         END_STRUCT;
         Reserve_5 : Struct
            ER_465 : Bool;   // Reserve
            ER_466 : Bool;   // Reserve
            ER_467 : Bool;   // Reserve
            ER_468 : Bool;   // Reserve
            ER_469 : Bool;   // Reserve
            ER_470 : Bool;   // Reserve
            ER_471 : Bool;   // Reserve
            ER_472 : Bool;   // Reserve
            ER_473 : Bool;   // Reserve
            ER_474 : Bool;   // Reserve
            ER_475 : Bool;   // Reserve
            ER_476 : Bool;   // Reserve
            ER_477 : Bool;   // Reserve
            ER_478 : Bool;   // Reserve
            ER_479 : Bool;   // Reserve
            ER_480 : Bool;   // Reserve
         END_STRUCT;
         Reserve_6 : Struct   // Meldungen Reserve
            ER_301 : Bool;   // Reserve
            ER_302 : Bool;   // Reserve
            ER_303 : Bool;   // Reserve
            ER_304 : Bool;   // Reserve
            ER_305 : Bool;   // Reserve
            ER_306 : Bool;   // Reserve
            ER_307 : Bool;   // Reserve
            ER_308 : Bool;   // Reserve
            ER_309 : Bool;   // Reserve
            ER_310 : Bool;   // Reserve
            ER_311 : Bool;   // Reserve
            ER_312 : Bool;   // Reserve
            ER_313 : Bool;   // Reserve
            ER_314 : Bool;   // Reserve
            ER_315 : Bool;   // Reserve
            ER_316 : Bool;   // Reserve
         END_STRUCT;
         Reserve_7 : Struct   // Meldungen Reserve
            ER_317 : Bool;   // Reserve
            ER_318 : Bool;   // Reserve
            ER_319 : Bool;   // Reserve
            ER_320 : Bool;   // Reserve
            ER_321 : Bool;   // Reserve
            ER_322 : Bool;   // Reserve
            ER_323 : Bool;   // Reserve
            ER_324 : Bool;   // Reserve
            ER_325 : Bool;   // Reserve
            ER_326 : Bool;   // Reserve
            ER_327 : Bool;   // Reserve
            ER_328 : Bool;   // Reserve
            ER_329 : Bool;   // Reserve
            ER_330 : Bool;   // Reserve
            ER_331 : Bool;   // Reserve
            ER_332 : Bool;   // Reserve
         END_STRUCT;
         Reserve_8 : Struct   // FU Reserve
            ER_333 : Bool;   // Störung Reserve FU 1: Überstrom
            ER_334 : Bool;   // Störung Reserve FU 1: Zwischenkreisspannung Überspannung
            ER_335 : Bool;   // Störung Reserve FU 1: Zwischenkreisspannung Unterspannung
            ER_336 : Bool;   // Störung Reserve FU 1: Übertemperatur Kühlkörper Wechselrichter
            ER_337 : Bool;   // Störung Reserve FU 1: Motordatenidentifikation fehlerhaft
            ER_338 : Bool;   // Störung Reserve FU 1: Erdschluss
            ER_339 : Bool;   // Störung Reserve FU 1: Reserve
            ER_340 : Bool;   // Störung Reserve FU 1: Führung durch PLC fehlt
            ER_341 : Bool;   // Störung Reserve FU 1: Reserve
            ER_342 : Bool;   // Störung Reserve FU 1: Reserve
            ER_343 : Bool;   // Störung Reserve FU 1: Reserve
            ER_344_ : Bool;   // Störung Reserve FU 1: Reserve
            ER_345 : Bool;   // Störung Reserve FU 1: Reserve
            ER_346 : Bool;   // Störung Reserve FU 1: Reserve
            ER_347 : Bool;   // Störung Reserve FU 1: Reserve
            ER_348 : Bool;   // Störung Reserve FU 1: Reserve
         END_STRUCT;
         Reserve_9 : Struct
            ER_349 : Bool;   // Reserve
            ER_350 : Bool;   // Reserve
            ER_351 : Bool;   // Reserve
            ER_352 : Bool;   // Reserve
            ER_353 : Bool;   // Reserve
            ER_354 : Bool;   // Reserve
            ER_355 : Bool;   // Reserve
            ER_356 : Bool;   // Reserve
            ER_357 : Bool;   // Reserve
            ER_358 : Bool;   // Reserve
            ER_359 : Bool;   // Reserve
            ER_360 : Bool;   // Reserve
            ER_361 : Bool;   // Reserve
            ER_362 : Bool;   // Reserve
            ER_363 : Bool;   // Reserve
            ER_364 : Bool;   // Reserve
         END_STRUCT;
         Reserve_10 : Struct   // FU Reserve
            ER_365 : Bool;   // Störung Reserve FU 2: Überstrom
            ER_366 : Bool;   // Störung Reserve FU 2: Zwischenkreisspannung Überspannung
            ER_367 : Bool;   // Störung Reserve FU 2: Zwischenkreisspannung Unterspannung
            ER_368 : Bool;   // Störung Reserve FU 2: Übertemperatur Kühlkörper Wechselrichter
            ER_369 : Bool;   // Störung Reserve FU 2: Motordatenidentifikation fehlerhaft
            ER_370 : Bool;   // Störung Reserve FU 2: Erdschluss
            ER_371 : Bool;   // Störung Reserve FU 2: Reserve
            ER_372 : Bool;   // Störung Reserve FU 2: Führung durch PLC fehlt
            ER_373 : Bool;   // Störung Reserve FU 2: Reserve
            ER_374 : Bool;   // Störung Reserve FU 2: Reserve
            ER_375 : Bool;   // Störung Reserve FU 2: Reserve
            ER_376 : Bool;   // Störung Reserve FU 2: Reserve
            ER_377 : Bool;   // Störung Reserve FU 2: Reserve
            ER_378 : Bool;   // Störung Reserve FU 2: Reserve
            ER_379 : Bool;   // Störung Reserve FU 2: Reserve
            ER_380 : Bool;   // Störung Reserve FU 2: Reserve
         END_STRUCT;
         SDC : Struct   // SDC Störungs
            ER_901 : Bool;   // Reserve
            ER_902 : Bool;   // Reserve
            ER_903 : Bool;   // Störung SDC Positionssprung
            ER_904 : Bool;   // Störung SDC keine Sektion gefunden
            ER_905 : Bool;   // Störung SDC Kommandos nicht plausibel
            ER_906 : Bool;   // Störung SDC Positionsgrenzen
            ER_907 : Bool;   // Störung SDC falsche EMS Nummer
            ER_908 : Bool;   // Störung SDC falsche Sektion Nummer
            ER_909 : Bool;   // Reserve
            ER_910 : Bool;   // Reserve
            ER_911 : Bool;   // Reserve
            ER_912 : Bool;   // Reserve
            ER_913 : Bool;   // Reserve
            ER_914 : Bool;   // Reserve
            ER_915 : Bool;   // Reserve
            ER_916 : Bool;   // Reserve
         END_STRUCT;
      END_STRUCT;
      EMS_ER_WORDs : Array[1..200] of Struct   // EMS Störung WORDs
         ER_WORD : Array[0..24] of Word;   // Störworte
      END_STRUCT;
      SDC : Struct
         ER_917 : Bool;   // Störung SDC Kommunikation mit Anlagensteuerung
         ER_918 : Bool;   // Störung SDC Safety Kommunikation mit Anlagensteuerung
         ER_919 : Bool;   // Störung SDC Reserve
         ER_920 : Bool;   // Störung SDC Reserve
         ER_921 : Bool;   // Störung SDC Reserve
         ER_922 : Bool;   // Störung SDC Reserve
         ER_923 : Bool;   // Störung SDC Reserve
         ER_924 : Bool;   // Störung SDC Reserve
         ER_925 : Bool;   // Störung SDC OB80 Zykluszeit
         ER_926 : Bool;   // Störung SDC OB82 Diagnosealarm
         ER_927 : Bool;   // Störung SDC OB83 Baugruppenwechsel
         ER_928 : Bool;   // Störung SDC OB86 Baugruppenträger ausgefallen
         ER_929 : Bool;   // Störung SDC OB121 Programmierfehler
         ER_930 : Bool;   // Störung SDC OB122 Peripherie-Zugriff
         ER_931 : Bool;   // Störung SDC Reserve
         ER_932 : Bool;   // Störung SDC Reserve
      END_STRUCT;
   END_VAR
BEGIN
END_DATA_BLOCK

DATA_BLOCK "DB_SDC_ERRORS_STAT"   // DB3724
{ S7_Optimized_Access := 'FALSE' }
VERSION : 0.1
   VAR
      HEADER : Struct   // Struktur für Datenheader // nicht verschieben
         DB_NR : Int := 3724;   // DB Nummer
         MIN_NR_FAULT_STAT : Int := 1;   // Niedrigste Fehler Nummer im Daten DB
         MAX_NR_FAULT_STAT : Int := 200;   // Höchste Fehler Nummer im Daten DB
         START_FAULT_STAT : Int := 20;   // Startadresse der Fehler Daten im Daten DB
         LAENGE_FAULT_STAT : Int := 28;   // Länge Fehler Daten
         FAULT_PRO_SEITE_HMI : Int := 10;   // Reserve
         RES12 : Int := 0;   // Reserve
         RES14 : Int := 0;   // Reserve
         RES16 : Int := 0;   // Reserve
         LOAD : Bool := FALSE;   // "0" zum laden des DB auf CPU
         RESET_ARCH : Bool := FALSE;   // Archiv löschen
      END_STRUCT;
      ER_ARCHIV : Array[1..1000] of "UDT_SDC_ERROR_STAT";   // Error Archiv
      ER_AKT : Array[1..200] of Struct   // Error aktiv EMS
         ER_TRIGER : Word;   // Error auslösen Aktiv von EMS
         ER_STAT : Array[1..4] of "UDT_SDC_TS_IF_STATUS_VAL";   // Error Status Aktiv EMS
      END_STRUCT;
   END_VAR
BEGIN
   ER_ARCHIV[1].EMS_TS_STAT_VAL.EMS_ID := 0;
   ER_ARCHIV[1].EMS_TS_STAT_VAL.PROFIL := 0;
   ER_ARCHIV[1].EMS_TS_STAT_VAL.DRIVE_POS := 0;
   ER_ARCHIV[1].EMS_TS_STAT_VAL.HOIST_POS := 0;
   ER_ARCHIV[1].EMS_TS_STAT_VAL.ERROR := 0;
   ER_ARCHIV[1].EMS_TS_STAT_VAL.DRIVE_POS_PERC := 0;
   ER_ARCHIV[1].EMS_TS_STAT_VAL.SEK := 0;
   ER_ARCHIV[1].ER._901_ER_SUM := FALSE;
   ER_ARCHIV[1].ER._902_ER_SUM_SDC := FALSE;
   ER_ARCHIV[1].ER._903_ER_BC_JUMP := FALSE;
   ER_ARCHIV[1].ER._904_ER_NO_SEK := FALSE;
   ER_ARCHIV[1].ER._905_ER_COMMAND := FALSE;
   ER_ARCHIV[1].ER._906_ER_BC_LIM := FALSE;
   ER_ARCHIV[1].ER._907_ER_EMS_ID := FALSE;
   ER_ARCHIV[1].ER._908_ER_SEK_NR := FALSE;
   ER_ARCHIV[1].ER._909_ER_LIFE := FALSE;
   ER_ARCHIV[1].ER._910_ER_BUS := FALSE;
   ER_ARCHIV[1].ER._911 := FALSE;
   ER_ARCHIV[1].ER._912 := FALSE;
   ER_ARCHIV[1].ER._913 := FALSE;
   ER_ARCHIV[1].ER._914 := FALSE;
   ER_ARCHIV[1].ER._915 := FALSE;
   ER_ARCHIV[1].ER._916 := FALSE;
   ER_ARCHIV[1].Spare := 0;
   ER_ARCHIV[1].ER_DATE := DT#1990-01-01-00:00:00;
   ER_ARCHIV[2].EMS_TS_STAT_VAL.EMS_ID := 0;
   ER_ARCHIV[2].EMS_TS_STAT_VAL.PROFIL := 0;
   ER_ARCHIV[2].EMS_TS_STAT_VAL.DRIVE_POS := 0;
   ER_ARCHIV[2].EMS_TS_STAT_VAL.HOIST_POS := 0;
   ER_ARCHIV[2].EMS_TS_STAT_VAL.ERROR := 0;
   ER_ARCHIV[2].EMS_TS_STAT_VAL.DRIVE_POS_PERC := 0;
   ER_ARCHIV[2].EMS_TS_STAT_VAL.SEK := 0;
   ER_ARCHIV[2].ER._901_ER_SUM := FALSE;
   ER_ARCHIV[2].ER._902_ER_SUM_SDC := FALSE;
   ER_ARCHIV[2].ER._903_ER_BC_JUMP := FALSE;
   ER_ARCHIV[2].ER._904_ER_NO_SEK := FALSE;
   ER_ARCHIV[2].ER._905_ER_COMMAND := FALSE;
   ER_ARCHIV[2].ER._906_ER_BC_LIM := FALSE;
   ER_ARCHIV[2].ER._907_ER_EMS_ID := FALSE;
   ER_ARCHIV[2].ER._908_ER_SEK_NR := FALSE;
   ER_ARCHIV[2].ER._909_ER_LIFE := FALSE;
   ER_ARCHIV[2].ER._910_ER_BUS := FALSE;
   ER_ARCHIV[2].ER._911 := FALSE;
   ER_ARCHIV[2].ER._912 := FALSE;
   ER_ARCHIV[2].ER._913 := FALSE;
   ER_ARCHIV[2].ER._914 := FALSE;
   ER_ARCHIV[2].ER._915 := FALSE;
   ER_ARCHIV[2].ER._916 := FALSE;
   ER_ARCHIV[2].Spare := 0;
   ER_ARCHIV[2].ER_DATE := DT#1990-01-01-00:00:00;
   ER_ARCHIV[3].EMS_TS_STAT_VAL.EMS_ID := 0;
   ER_ARCHIV[3].EMS_TS_STAT_VAL.PROFIL := 0;
   ER_ARCHIV[3].EMS_TS_STAT_VAL.DRIVE_POS := 0;
   ER_ARCHIV[3].EMS_TS_STAT_VAL.HOIST_POS := 0;
   ER_ARCHIV[3].EMS_TS_STAT_VAL.ERROR := 0;
   ER_ARCHIV[3].EMS_TS_STAT_VAL.DRIVE_POS_PERC := 0;
   ER_ARCHIV[3].EMS_TS_STAT_VAL.SEK := 0;
   ER_ARCHIV[3].ER._901_ER_SUM := FALSE;
   ER_ARCHIV[3].ER._902_ER_SUM_SDC := FALSE;
   ER_ARCHIV[3].ER._903_ER_BC_JUMP := FALSE;
   ER_ARCHIV[3].ER._904_ER_NO_SEK := FALSE;
   ER_ARCHIV[3].ER._905_ER_COMMAND := FALSE;
   ER_ARCHIV[3].ER._906_ER_BC_LIM := FALSE;
   ER_ARCHIV[3].ER._907_ER_EMS_ID := FALSE;
   ER_ARCHIV[3].ER._908_ER_SEK_NR := FALSE;
   ER_ARCHIV[3].ER._909_ER_LIFE := FALSE;
   ER_ARCHIV[3].ER._910_ER_BUS := FALSE;
   ER_ARCHIV[3].ER._911 := FALSE;
   ER_ARCHIV[3].ER._912 := FALSE;
   ER_ARCHIV[3].ER._913 := FALSE;
   ER_ARCHIV[3].ER._914 := FALSE;
   ER_ARCHIV[3].ER._915 := FALSE;
   ER_ARCHIV[3].ER._916 := FALSE;
   ER_ARCHIV[3].Spare := 0;
   ER_ARCHIV[3].ER_DATE := DT#1990-01-01-00:00:00;
   ER_ARCHIV[4].EMS_TS_STAT_VAL.EMS_ID := 0;
   ER_ARCHIV[4].EMS_TS_STAT_VAL.PROFIL := 0;
   ER_ARCHIV[4].EMS_TS_STAT_VAL.DRIVE_POS := 0;
   ER_ARCHIV[4].EMS_TS_STAT_VAL.HOIST_POS := 0;
   ER_ARCHIV[4].EMS_TS_STAT_VAL.ERROR := 0;
   ER_ARCHIV[4].EMS_TS_STAT_VAL.DRIVE_POS_PERC := 0;
   ER_ARCHIV[4].EMS_TS_STAT_VAL.SEK := 0;
   ER_ARCHIV[4].ER._901_ER_SUM := FALSE;
   ER_ARCHIV[4].ER._902_ER_SUM_SDC := FALSE;
   ER_ARCHIV[4].ER._903_ER_BC_JUMP := FALSE;
   ER_ARCHIV[4].ER._904_ER_NO_SEK := FALSE;
   ER_ARCHIV[4].ER._905_ER_COMMAND := FALSE;
   ER_ARCHIV[4].ER._906_ER_BC_LIM := FALSE;
   ER_ARCHIV[4].ER._907_ER_EMS_ID := FALSE;
   ER_ARCHIV[4].ER._908_ER_SEK_NR := FALSE;
   ER_ARCHIV[4].ER._909_ER_LIFE := FALSE;
   ER_ARCHIV[4].ER._910_ER_BUS := FALSE;
   ER_ARCHIV[4].ER._911 := FALSE;
   ER_ARCHIV[4].ER._912 := FALSE;
   ER_ARCHIV[4].ER._913 := FALSE;
   ER_ARCHIV[4].ER._914 := FALSE;
   ER_ARCHIV[4].ER._915 := FALSE;
   ER_ARCHIV[4].ER._916 := FALSE;
   ER_ARCHIV[4].Spare := 0;
   ER_ARCHIV[4].ER_DATE := DT#1990-01-01-00:00:00;
   ER_ARCHIV[5].EMS_TS_STAT_VAL.EMS_ID := 0;
   ER_ARCHIV[5].EMS_TS_STAT_VAL.PROFIL := 0;
   ER_ARCHIV[5].EMS_TS_STAT_VAL.DRIVE_POS := 0;
   ER_ARCHIV[5].EMS_TS_STAT_VAL.HOIST_POS := 0;
   ER_ARCHIV[5].EMS_TS_STAT_VAL.ERROR := 0;
   ER_ARCHIV[5].EMS_TS_STAT_VAL.DRIVE_POS_PERC := 0;
   ER_ARCHIV[5].EMS_TS_STAT_VAL.SEK := 0;
   ER_ARCHIV[5].ER._901_ER_SUM := FALSE;
   ER_ARCHIV[5].ER._902_ER_SUM_SDC := FALSE;
   ER_ARCHIV[5].ER._903_ER_BC_JUMP := FALSE;
   ER_ARCHIV[5].ER._904_ER_NO_SEK := FALSE;
   ER_ARCHIV[5].ER._905_ER_COMMAND := FALSE;
   ER_ARCHIV[5].ER._906_ER_BC_LIM := FALSE;
   ER_ARCHIV[5].ER._907_ER_EMS_ID := FALSE;
   ER_ARCHIV[5].ER._908_ER_SEK_NR := FALSE;
   ER_ARCHIV[5].ER._909_ER_LIFE := FALSE;
   ER_ARCHIV[5].ER._910_ER_BUS := FALSE;
   ER_ARCHIV[5].ER._911 := FALSE;
   ER_ARCHIV[5].ER._912 := FALSE;
   ER_ARCHIV[5].ER._913 := FALSE;
   ER_ARCHIV[5].ER._914 := FALSE;
   ER_ARCHIV[5].ER._915 := FALSE;
   ER_ARCHIV[5].ER._916 := FALSE;
   ER_ARCHIV[5].Spare := 0;
   ER_ARCHIV[5].ER_DATE := DT#1990-01-01-00:00:00;
   ER_ARCHIV[6].EMS_TS_STAT_VAL.EMS_ID := 0;
   ER_ARCHIV[6].EMS_TS_STAT_VAL.PROFIL := 0;
   ER_ARCHIV[6].EMS_TS_STAT_VAL.DRIVE_POS := 0;
   ER_ARCHIV[6].EMS_TS_STAT_VAL.HOIST_POS := 0;
   ER_ARCHIV[6].EMS_TS_STAT_VAL.ERROR := 0;
   ER_ARCHIV[6].EMS_TS_STAT_VAL.DRIVE_POS_PERC := 0;
   ER_ARCHIV[6].EMS_TS_STAT_VAL.SEK := 0;
   ER_ARCHIV[6].ER._901_ER_SUM := FALSE;
   ER_ARCHIV[6].ER._902_ER_SUM_SDC := FALSE;
   ER_ARCHIV[6].ER._903_ER_BC_JUMP := FALSE;
   ER_ARCHIV[6].ER._904_ER_NO_SEK := FALSE;
   ER_ARCHIV[6].ER._905_ER_COMMAND := FALSE;
   ER_ARCHIV[6].ER._906_ER_BC_LIM := FALSE;
   ER_ARCHIV[6].ER._907_ER_EMS_ID := FALSE;
   ER_ARCHIV[6].ER._908_ER_SEK_NR := FALSE;
   ER_ARCHIV[6].ER._909_ER_LIFE := FALSE;
   ER_ARCHIV[6].ER._910_ER_BUS := FALSE;
   ER_ARCHIV[6].ER._911 := FALSE;
   ER_ARCHIV[6].ER._912 := FALSE;
   ER_ARCHIV[6].ER._913 := FALSE;
   ER_ARCHIV[6].ER._914 := FALSE;
   ER_ARCHIV[6].ER._915 := FALSE;
   ER_ARCHIV[6].ER._916 := FALSE;
   ER_ARCHIV[6].Spare := 0;
   ER_ARCHIV[6].ER_DATE := DT#1990-01-01-00:00:00;
   ER_ARCHIV[7].EMS_TS_STAT_VAL.EMS_ID := 0;
   ER_ARCHIV[7].EMS_TS_STAT_VAL.PROFIL := 0;
   ER_ARCHIV[7].EMS_TS_STAT_VAL.DRIVE_POS := 0;
   ER_ARCHIV[7].EMS_TS_STAT_VAL.HOIST_POS := 0;
   ER_ARCHIV[7].EMS_TS_STAT_VAL.ERROR := 0;
   ER_ARCHIV[7].EMS_TS_STAT_VAL.DRIVE_POS_PERC := 0;
   ER_ARCHIV[7].EMS_TS_STAT_VAL.SEK := 0;
   ER_ARCHIV[7].ER._901_ER_SUM := FALSE;
   ER_ARCHIV[7].ER._902_ER_SUM_SDC := FALSE;
   ER_ARCHIV[7].ER._903_ER_BC_JUMP := FALSE;
   ER_ARCHIV[7].ER._904_ER_NO_SEK := FALSE;
   ER_ARCHIV[7].ER._905_ER_COMMAND := FALSE;
   ER_ARCHIV[7].ER._906_ER_BC_LIM := FALSE;
   ER_ARCHIV[7].ER._907_ER_EMS_ID := FALSE;
   ER_ARCHIV[7].ER._908_ER_SEK_NR := FALSE;
   ER_ARCHIV[7].ER._909_ER_LIFE := FALSE;
   ER_ARCHIV[7].ER._910_ER_BUS := FALSE;
   ER_ARCHIV[7].ER._911 := FALSE;
   ER_ARCHIV[7].ER._912 := FALSE;
   ER_ARCHIV[7].ER._913 := FALSE;
   ER_ARCHIV[7].ER._914 := FALSE;
   ER_ARCHIV[7].ER._915 := FALSE;
   ER_ARCHIV[7].ER._916 := FALSE;
   ER_ARCHIV[7].Spare := 0;
   ER_ARCHIV[7].ER_DATE := DT#1990-01-01-00:00:00;
   ER_ARCHIV[8].EMS_TS_STAT_VAL.EMS_ID := 0;
   ER_ARCHIV[8].EMS_TS_STAT_VAL.PROFIL := 0;
   ER_ARCHIV[8].EMS_TS_STAT_VAL.DRIVE_POS := 0;
   ER_ARCHIV[8].EMS_TS_STAT_VAL.HOIST_POS := 0;
   ER_ARCHIV[8].EMS_TS_STAT_VAL.ERROR := 0;
   ER_ARCHIV[8].EMS_TS_STAT_VAL.DRIVE_POS_PERC := 0;
   ER_ARCHIV[8].EMS_TS_STAT_VAL.SEK := 0;
   ER_ARCHIV[8].ER._901_ER_SUM := FALSE;
   ER_ARCHIV[8].ER._902_ER_SUM_SDC := FALSE;
   ER_ARCHIV[8].ER._903_ER_BC_JUMP := FALSE;
   ER_ARCHIV[8].ER._904_ER_NO_SEK := FALSE;
   ER_ARCHIV[8].ER._905_ER_COMMAND := FALSE;
   ER_ARCHIV[8].ER._906_ER_BC_LIM := FALSE;
   ER_ARCHIV[8].ER._907_ER_EMS_ID := FALSE;
   ER_ARCHIV[8].ER._908_ER_SEK_NR := FALSE;
   ER_ARCHIV[8].ER._909_ER_LIFE := FALSE;
   ER_ARCHIV[8].ER._910_ER_BUS := FALSE;
   ER_ARCHIV[8].ER._911 := FALSE;
   ER_ARCHIV[8].ER._912 := FALSE;
   ER_ARCHIV[8].ER._913 := FALSE;
   ER_ARCHIV[8].ER._914 := FALSE;
   ER_ARCHIV[8].ER._915 := FALSE;
   ER_ARCHIV[8].ER._916 := FALSE;
   ER_ARCHIV[8].Spare := 0;
   ER_ARCHIV[8].ER_DATE := DT#1990-01-01-00:00:00;
   // 30600 more start values not shown
END_DATA_BLOCK

DATA_BLOCK "DB_SDC_EMS_SIM"   // DB3726
{ S7_Optimized_Access := 'FALSE' }
VERSION : 0.1
   VAR
      HEADER : Struct   // Struktur für Datenheader // nicht verschieben
         DB_NR : Int := 3726;   // DB Nummer
         MIN_NR_EMS : Int := 1;   // Niedrigste EMS Nummer im Daten DB
         MAX_NR_EMS : Int := 200;   // Höchste EMS Nummer im Daten DB
         START_DAT : Int := 40;   // Startadresse der EMS Daten im Daten DB
         LAENGE_EMS : Int := 40;   // Länge Eingänge pro EMS
         RES10 : Int := 0;   // Reserve
         RES12 : Int := 0;   // Reserve
         RES14 : Int := 0;   // Reserve
         RES16 : Int := 0;   // Reserve
         RES18 : Int := 0;   // Reserve
      END_STRUCT;
      PAR : Struct   // Parameter Simulation
         BARCODE_START : DInt := 1;   // min Barcodevalue
         BARCODE_ENDE : DInt := 500000;   // max Barcodevalue
         HUB_START : Int := 0;   // min Hoistvalue
         HUB_ENDE : Int := 4010;   // max Hoistvalue
         LEAP_AKT : Array[1..20] of Bool;   // Leap Aktiv
         LEAP_HIGH_LOW : Array[1..20] of Bool;   // Leap Aktiv
         ON : Bool := TRUE;   // Simulation ON "1"
         RES18 : Int := 0;   // Reserve
      END_STRUCT;
      EMS : Array[1..200] of "UDT_EMS_IF_Q";   // EMS Simulation Eingänge
      EMS_TEMP : "UDT_EMS_IF_Q";
   END_VAR
BEGIN
   PAR.LEAP_AKT[1] := TRUE;
   PAR.LEAP_AKT[2] := TRUE;
   PAR.LEAP_AKT[3] := TRUE;
   PAR.LEAP_HIGH_LOW[1] := TRUE;
   PAR.LEAP_HIGH_LOW[2] := FALSE;
   PAR.LEAP_HIGH_LOW[3] := TRUE;
   PAR.LEAP_AKT[4] := FALSE;
   PAR.LEAP_AKT[5] := FALSE;
   PAR.LEAP_AKT[6] := FALSE;
   PAR.LEAP_AKT[7] := FALSE;
   PAR.LEAP_AKT[8] := FALSE;
   PAR.LEAP_AKT[9] := FALSE;
   PAR.LEAP_AKT[10] := FALSE;
   PAR.LEAP_AKT[11] := FALSE;
   PAR.LEAP_AKT[12] := FALSE;
   PAR.LEAP_AKT[13] := FALSE;
   PAR.LEAP_AKT[14] := FALSE;
   PAR.LEAP_AKT[15] := FALSE;
   PAR.LEAP_AKT[16] := FALSE;
   PAR.LEAP_AKT[17] := FALSE;
   PAR.LEAP_AKT[18] := FALSE;
   PAR.LEAP_AKT[19] := FALSE;
   PAR.LEAP_AKT[20] := FALSE;
   PAR.LEAP_HIGH_LOW[4] := FALSE;
   PAR.LEAP_HIGH_LOW[5] := FALSE;
   PAR.LEAP_HIGH_LOW[6] := FALSE;
   PAR.LEAP_HIGH_LOW[7] := FALSE;
   PAR.LEAP_HIGH_LOW[8] := FALSE;
   PAR.LEAP_HIGH_LOW[9] := FALSE;
   PAR.LEAP_HIGH_LOW[10] := FALSE;
   PAR.LEAP_HIGH_LOW[11] := FALSE;
   PAR.LEAP_HIGH_LOW[12] := FALSE;
   PAR.LEAP_HIGH_LOW[13] := FALSE;
   PAR.LEAP_HIGH_LOW[14] := FALSE;
   PAR.LEAP_HIGH_LOW[15] := FALSE;
   PAR.LEAP_HIGH_LOW[16] := FALSE;
   PAR.LEAP_HIGH_LOW[17] := FALSE;
   PAR.LEAP_HIGH_LOW[18] := FALSE;
   PAR.LEAP_HIGH_LOW[19] := FALSE;
   PAR.LEAP_HIGH_LOW[20] := FALSE;
   EMS[1].STAT.LIFE_BIT := TRUE;
   EMS[1].STAT.ER_SUM := FALSE;
   EMS[1].STAT.IR_MAN := FALSE;
   EMS[1].STAT.ER_RESET := FALSE;
   EMS[1].STAT.HOIST_CLEAR := FALSE;
   EMS[1].STAT.POS_START_X := FALSE;
   EMS[1].STAT.ALWAYS_ONE := TRUE;
   EMS[1].STAT.H_DISABLED := FALSE;
   EMS[1].STAT.D_FWD := TRUE;
   EMS[1].STAT.D_RWD := FALSE;
   EMS[1].STAT.bit12 := FALSE;
   EMS[1].STAT.D_IN_POS := FALSE;
   EMS[1].STAT.H_UP := FALSE;
   EMS[1].STAT.H_DOWN := FALSE;
   EMS[1].STAT.H_IN_POS := TRUE;
   EMS[1].STAT.H_IN_TOPPOS := FALSE;
   EMS[1].STAT.bit2_0 := FALSE;
   EMS[1].STAT.bit2_1 := FALSE;
   EMS[1].STAT.bit2_2 := FALSE;
   EMS[1].STAT.bit2_3 := FALSE;
   EMS[1].STAT.IN_BOTPOS := FALSE;
   EMS[1].STAT.bit2_5 := FALSE;
   EMS[1].STAT.bit2_6 := FALSE;
   EMS[1].STAT.bit2_7 := FALSE;
   EMS[1].STAT.MESS_POS := FALSE;
   EMS[1].STAT.bit3_2 := FALSE;
   EMS[1].STAT.bit3_3 := FALSE;
   EMS[1].STAT.bit3_4 := FALSE;
   EMS[1].STAT.bit3_5 := FALSE;
   EMS[1].STAT.bit3_6 := FALSE;
   EMS[1].STAT.DATA_TRANS := FALSE;
   EMS[1].ERROR := 0;
   EMS[1].D_POS := 22899;
   EMS[1].H_POS := 603;
   EMS[1].ER_WORD_No := 1;
   EMS[1].ER_WORD := 16#0000;
   EMS[1].FB_DBNo := 0;
   EMS[1].FB_DBBNo := 0;
   EMS[2].STAT.LIFE_BIT := TRUE;
   EMS[2].STAT.ER_SUM := FALSE;
   EMS[2].STAT.IR_MAN := FALSE;
   EMS[2].STAT.ER_RESET := FALSE;
   EMS[2].STAT.HOIST_CLEAR := FALSE;
   EMS[2].STAT.POS_START_X := FALSE;
   EMS[2].STAT.ALWAYS_ONE := TRUE;
   EMS[2].STAT.H_DISABLED := FALSE;
   EMS[2].STAT.D_FWD := TRUE;
   EMS[2].STAT.D_RWD := FALSE;
   EMS[2].STAT.bit12 := FALSE;
   EMS[2].STAT.D_IN_POS := FALSE;
   EMS[2].STAT.H_UP := FALSE;
   EMS[2].STAT.H_DOWN := FALSE;
   EMS[2].STAT.H_IN_POS := FALSE;
   EMS[2].STAT.H_IN_TOPPOS := TRUE;
   EMS[2].STAT.bit2_0 := FALSE;
   EMS[2].STAT.bit2_1 := FALSE;
   EMS[2].STAT.bit2_2 := FALSE;
   EMS[2].STAT.bit2_3 := FALSE;
   EMS[2].STAT.IN_BOTPOS := FALSE;
   EMS[2].STAT.bit2_5 := FALSE;
   EMS[2].STAT.bit2_6 := FALSE;
   EMS[2].STAT.bit2_7 := FALSE;
   EMS[2].STAT.MESS_POS := FALSE;
   EMS[2].STAT.bit3_2 := FALSE;
   EMS[2].STAT.bit3_3 := FALSE;
   EMS[2].STAT.bit3_4 := FALSE;
   EMS[2].STAT.bit3_5 := FALSE;
   EMS[2].STAT.bit3_6 := FALSE;
   EMS[2].STAT.DATA_TRANS := FALSE;
   EMS[2].ERROR := 0;
   EMS[2].D_POS := 10522;
   EMS[2].H_POS := 4010;
   EMS[2].ER_WORD_No := 1;
   EMS[2].ER_WORD := 16#0000;
   EMS[2].FB_DBNo := 0;
   EMS[2].FB_DBBNo := 0;
   EMS[3].STAT.LIFE_BIT := TRUE;
   EMS[3].STAT.ER_SUM := FALSE;
   EMS[3].STAT.IR_MAN := FALSE;
   EMS[3].STAT.ER_RESET := FALSE;
   EMS[3].STAT.HOIST_CLEAR := FALSE;
   EMS[3].STAT.POS_START_X := FALSE;
   EMS[3].STAT.ALWAYS_ONE := TRUE;
   EMS[3].STAT.H_DISABLED := FALSE;
   EMS[3].STAT.D_FWD := TRUE;
   EMS[3].STAT.D_RWD := FALSE;
   EMS[3].STAT.bit12 := FALSE;
   EMS[3].STAT.D_IN_POS := FALSE;
   EMS[3].STAT.H_UP := FALSE;
   EMS[3].STAT.H_DOWN := FALSE;
   EMS[3].STAT.H_IN_POS := FALSE;
   EMS[3].STAT.H_IN_TOPPOS := TRUE;
   EMS[3].STAT.bit2_0 := FALSE;
   EMS[3].STAT.bit2_1 := FALSE;
   EMS[3].STAT.bit2_2 := FALSE;
   EMS[3].STAT.bit2_3 := FALSE;
   EMS[3].STAT.IN_BOTPOS := FALSE;
   EMS[3].STAT.bit2_5 := FALSE;
   EMS[3].STAT.bit2_6 := FALSE;
   EMS[3].STAT.bit2_7 := FALSE;
   EMS[3].STAT.MESS_POS := FALSE;
   EMS[3].STAT.bit3_2 := FALSE;
   EMS[3].STAT.bit3_3 := FALSE;
   EMS[3].STAT.bit3_4 := FALSE;
   EMS[3].STAT.bit3_5 := FALSE;
   EMS[3].STAT.bit3_6 := FALSE;
   EMS[3].STAT.DATA_TRANS := FALSE;
   EMS[3].ERROR := 0;
   EMS[3].D_POS := 96650;
   EMS[3].H_POS := 4010;
   EMS[3].ER_WORD_No := 1;
   EMS[3].ER_WORD := 16#0000;
   EMS[3].FB_DBNo := 0;
   EMS[3].FB_DBBNo := 0;
   EMS[4].STAT.LIFE_BIT := FALSE;
   EMS[4].STAT.ER_SUM := FALSE;
   EMS[4].STAT.IR_MAN := FALSE;
   EMS[4].STAT.ER_RESET := FALSE;
   EMS[4].STAT.HOIST_CLEAR := FALSE;
   EMS[4].STAT.POS_START_X := FALSE;
   EMS[4].STAT.ALWAYS_ONE := FALSE;
   EMS[4].STAT.H_DISABLED := FALSE;
   EMS[4].STAT.D_FWD := FALSE;
   EMS[4].STAT.D_RWD := FALSE;
   EMS[4].STAT.bit12 := FALSE;
   EMS[4].STAT.D_IN_POS := FALSE;
   EMS[4].STAT.H_UP := FALSE;
   EMS[4].STAT.H_DOWN := FALSE;
   EMS[4].STAT.H_IN_POS := FALSE;
   EMS[4].STAT.H_IN_TOPPOS := FALSE;
   EMS[4].STAT.bit2_0 := FALSE;
   EMS[4].STAT.bit2_1 := FALSE;
   EMS[4].STAT.bit2_2 := FALSE;
   EMS[4].STAT.bit2_3 := FALSE;
   EMS[4].STAT.IN_BOTPOS := FALSE;
   EMS[4].STAT.bit2_5 := FALSE;
   EMS[4].STAT.bit2_6 := FALSE;
   EMS[4].STAT.bit2_7 := FALSE;
   EMS[4].STAT.MESS_POS := FALSE;
   EMS[4].STAT.bit3_2 := FALSE;
   EMS[4].STAT.bit3_3 := FALSE;
   EMS[4].STAT.bit3_4 := FALSE;
   EMS[4].STAT.bit3_5 := FALSE;
   EMS[4].STAT.bit3_6 := FALSE;
   EMS[4].STAT.DATA_TRANS := FALSE;
   EMS[4].ERROR := 0;
   EMS[4].D_POS := 0;
   EMS[4].H_POS := 0;
   EMS[4].ER_WORD_No := 0;
   EMS[4].ER_WORD := 16#0000;
   EMS[4].FB_DBNo := 0;
   EMS[4].FB_DBBNo := 0;
   EMS[5].STAT.LIFE_BIT := FALSE;
   EMS[5].STAT.ER_SUM := FALSE;
   EMS[5].STAT.IR_MAN := FALSE;
   EMS[5].STAT.ER_RESET := FALSE;
   EMS[5].STAT.HOIST_CLEAR := FALSE;
   EMS[5].STAT.POS_START_X := FALSE;
   EMS[5].STAT.ALWAYS_ONE := FALSE;
   EMS[5].STAT.H_DISABLED := FALSE;
   // 15719 more start values not shown
END_DATA_BLOCK

DATA_BLOCK "DB_SDC_EMS_TA"   // DB3728
{ S7_Optimized_Access := 'FALSE' }
VERSION : 0.1
   VAR
      HEADER : Struct
         DB_NR : Int := 3728;
         MIN_NR_EMS : Int := 1;
         MAX_NR_EMS : Int := 200;
         START_EMS : Int := 20;
         LAENGE_TA_DATA : Int := 6;
         ANZ_TA : Int := 3;
         Res120 : Int;
         Res140 : Int;
         Res160 : Int;
         Load : Bool := TRUE;
      END_STRUCT;
      EMS : Array[1..200] of Struct
         TA : Array[1..3] of "UDT_EMS_TA";
      END_STRUCT;
   END_VAR
BEGIN
END_DATA_BLOCK

DATA_BLOCK "DB_SDC_BARCODE_INSERTS"   // DB3734
{ S7_Optimized_Access := 'FALSE' }
VERSION : 0.1
   VAR
      HYST : Int := 100;   // Hysterese für Positionswerte
      INSERTS : Int := 2;   // Positioning Leaps
      INSERT : Array[1..20] of Struct   // LEAPs
         COURSELOW : DInt;   // lower position value Course Barocdevalue befor Insert
         COURSEHIGH : DInt;   // höhere Positionswert Course Barocde Wert nach Insert
         INSERTLOW : DInt;   // lower position value Barocdevalue Insert low
         INSERTHIGH : DInt;   // höhere Positionswert Barocde Wert liegt Hoch
         OFFSET : DInt;   // absoluten Offset zu Beginn der Einfügen -> zusätzlich von allen Einsätzen unter
      END_STRUCT;
      ABS_DIST_COURSE : DInt := 304270;   // abslolute Entfernung
   END_VAR
BEGIN
   INSERT[2].COURSELOW := 254280;
   INSERT[1].COURSEHIGH := 5800;
   INSERT[2].COURSEHIGH := 256410;
   INSERT[2].INSERTLOW := 0;
   INSERT[2].INSERTHIGH := 0;
   INSERT[1].OFFSET := -5800;
   INSERT[2].OFFSET := -7930;
   INSERT[1].COURSELOW := 0;
   INSERT[1].INSERTLOW := 0;
   INSERT[1].INSERTHIGH := 0;
   INSERT[3].COURSELOW := 0;
   INSERT[3].COURSEHIGH := 0;
   INSERT[3].INSERTLOW := 0;
   INSERT[3].INSERTHIGH := 0;
   INSERT[3].OFFSET := -1000;
   INSERT[4].COURSELOW := 0;
   INSERT[4].COURSEHIGH := 0;
   INSERT[4].INSERTLOW := 0;
   INSERT[4].INSERTHIGH := 0;
   INSERT[4].OFFSET := -1000;
   INSERT[5].COURSELOW := 0;
   INSERT[5].COURSEHIGH := 0;
   INSERT[5].INSERTLOW := 0;
   INSERT[5].INSERTHIGH := 0;
   INSERT[5].OFFSET := -1000;
   INSERT[6].COURSELOW := 0;
   INSERT[6].COURSEHIGH := 0;
   INSERT[6].INSERTLOW := 0;
   INSERT[6].INSERTHIGH := 0;
   INSERT[6].OFFSET := -1000;
   INSERT[7].COURSELOW := 0;
   INSERT[7].COURSEHIGH := 0;
   INSERT[7].INSERTLOW := 0;
   INSERT[7].INSERTHIGH := 0;
   INSERT[7].OFFSET := -1000;
   INSERT[8].COURSELOW := 0;
   INSERT[8].COURSEHIGH := 0;
   INSERT[8].INSERTLOW := 0;
   INSERT[8].INSERTHIGH := 0;
   INSERT[8].OFFSET := -1000;
   INSERT[9].COURSELOW := 0;
   INSERT[9].COURSEHIGH := 0;
   INSERT[9].INSERTLOW := 0;
   INSERT[9].INSERTHIGH := 0;
   INSERT[9].OFFSET := -1000;
   INSERT[10].COURSELOW := 0;
   INSERT[10].COURSEHIGH := 0;
   INSERT[10].INSERTLOW := 0;
   INSERT[10].INSERTHIGH := 0;
   INSERT[10].OFFSET := -1000;
   INSERT[11].COURSELOW := 0;
   INSERT[11].COURSEHIGH := 0;
   INSERT[11].INSERTLOW := 0;
   INSERT[11].INSERTHIGH := 0;
   INSERT[11].OFFSET := 0;
   INSERT[12].COURSELOW := 0;
   INSERT[12].COURSEHIGH := 0;
   INSERT[12].INSERTLOW := 0;
   INSERT[12].INSERTHIGH := 0;
   INSERT[12].OFFSET := 0;
   INSERT[13].COURSELOW := 0;
   INSERT[13].COURSEHIGH := 0;
   INSERT[13].INSERTLOW := 0;
   INSERT[13].INSERTHIGH := 0;
   INSERT[13].OFFSET := 0;
   INSERT[14].COURSELOW := 0;
   INSERT[14].COURSEHIGH := 0;
   INSERT[14].INSERTLOW := 0;
   INSERT[14].INSERTHIGH := 0;
   INSERT[14].OFFSET := 0;
   INSERT[15].COURSELOW := 0;
   INSERT[15].COURSEHIGH := 0;
   INSERT[15].INSERTLOW := 0;
   INSERT[15].INSERTHIGH := 0;
   INSERT[15].OFFSET := 0;
   INSERT[16].COURSELOW := 0;
   INSERT[16].COURSEHIGH := 0;
   INSERT[16].INSERTLOW := 0;
   INSERT[16].INSERTHIGH := 0;
   INSERT[16].OFFSET := 0;
   INSERT[17].COURSELOW := 0;
   INSERT[17].COURSEHIGH := 0;
   INSERT[17].INSERTLOW := 0;
   INSERT[17].INSERTHIGH := 0;
   INSERT[17].OFFSET := 0;
   INSERT[18].COURSELOW := 0;
   INSERT[18].COURSEHIGH := 0;
   INSERT[18].INSERTLOW := 0;
   INSERT[18].INSERTHIGH := 0;
   INSERT[18].OFFSET := 0;
   INSERT[19].COURSELOW := 0;
   INSERT[19].COURSEHIGH := 0;
   INSERT[19].INSERTLOW := 0;
   INSERT[19].INSERTHIGH := 0;
   INSERT[19].OFFSET := 0;
   INSERT[20].COURSELOW := 0;
   INSERT[20].COURSEHIGH := 0;
   INSERT[20].INSERTLOW := 0;
   INSERT[20].INSERTHIGH := 0;
   INSERT[20].OFFSET := 0;
END_DATA_BLOCK

DATA_BLOCK "DB_SDC_TS_REFERENCE_1"   // DB3780
{ S7_Optimized_Access := 'FALSE' }
VERSION : 0.1
   VAR
      HEADER : Struct
         DB_NR : Int := 3780;
         MIN_NR_SEK : Int := 1;
         MAX_NR_SEK : Int := 100;
         START_DAT : Int := 20;
         LAENGE_SEK_DATA : Int := 200;
         Res10 : Int := 0;
         Res12 : Int := 0;
         Res14 : Int := 0;
         Res16 : Int := 0;
         Res18 : Int := 0;
      END_STRUCT;
      Reference : Array[1..100] of Struct
         Sektion : Array[1..16] of Char;
         Actionpoint_1 : Array[1..16] of Char;
         Actionpoint_2 : Array[1..16] of Char;
         Height : Array[1..16] of Char;
         Hoist_offset_1 : Array[1..16] of Char;
         Hoist_offset_2 : Array[1..16] of Char;
         Hoist_offset_3 : Array[1..16] of Char;
         Hoist_offset_4 : Array[1..16] of Char;
         Reserve : Array[128..199] of Char;
      END_STRUCT;
   END_VAR
BEGIN
   Reference[1].Reserve[199] := ' ';
   Reference[1].Reserve[198] := ' ';
   Reference[1].Reserve[197] := ' ';
   Reference[1].Reserve[196] := ' ';
   Reference[1].Reserve[195] := ' ';
   Reference[1].Reserve[194] := ' ';
   Reference[1].Reserve[193] := ' ';
   Reference[1].Reserve[192] := ' ';
   Reference[1].Reserve[191] := ' ';
   Reference[1].Reserve[190] := ' ';
   Reference[1].Reserve[189] := ' ';
   Reference[1].Reserve[188] := ' ';
   Reference[1].Reserve[187] := ' ';
   Reference[1].Reserve[186] := ' ';
   Reference[1].Reserve[185] := ' ';
   Reference[1].Reserve[184] := ' ';
   Reference[1].Reserve[183] := ' ';
   Reference[1].Reserve[182] := ' ';
   Reference[1].Reserve[181] := ' ';
   Reference[1].Reserve[180] := ' ';
   Reference[1].Reserve[179] := ' ';
   Reference[1].Reserve[178] := ' ';
   Reference[1].Reserve[177] := ' ';
   Reference[1].Reserve[176] := ' ';
   Reference[1].Reserve[175] := ' ';
   Reference[1].Reserve[174] := ' ';
   Reference[1].Reserve[173] := ' ';
   Reference[1].Reserve[172] := ' ';
   Reference[1].Reserve[171] := ' ';
   Reference[1].Reserve[170] := ' ';
   Reference[1].Reserve[169] := ' ';
   Reference[1].Reserve[168] := ' ';
   Reference[1].Reserve[167] := ' ';
   Reference[1].Reserve[166] := ' ';
   Reference[1].Reserve[165] := ' ';
   Reference[1].Reserve[164] := ' ';
   Reference[1].Reserve[163] := ' ';
   Reference[1].Reserve[162] := ' ';
   Reference[1].Reserve[161] := ' ';
   Reference[1].Reserve[160] := ' ';
   Reference[1].Reserve[159] := ' ';
   Reference[1].Reserve[158] := ' ';
   Reference[1].Reserve[157] := ' ';
   Reference[1].Reserve[156] := ' ';
   Reference[1].Reserve[155] := ' ';
   Reference[1].Reserve[154] := ' ';
   Reference[1].Reserve[153] := ' ';
   Reference[1].Reserve[152] := ' ';
   Reference[1].Reserve[151] := ' ';
   Reference[1].Reserve[150] := ' ';
   Reference[1].Reserve[149] := ' ';
   Reference[1].Reserve[148] := ' ';
   Reference[1].Reserve[147] := ' ';
   Reference[1].Reserve[146] := ' ';
   Reference[1].Reserve[145] := ' ';
   Reference[1].Reserve[144] := ' ';
   Reference[1].Reserve[143] := '0';
   Reference[1].Reserve[142] := '0';
   Reference[1].Reserve[141] := '0';
   Reference[1].Reserve[140] := '0';
   Reference[1].Reserve[139] := '0';
   Reference[1].Reserve[138] := '0';
   Reference[1].Reserve[137] := '0';
   Reference[1].Reserve[136] := '0';
   Reference[1].Reserve[135] := '0';
   Reference[1].Reserve[134] := '0';
   Reference[1].Reserve[133] := '0';
   Reference[1].Reserve[132] := '0';
   Reference[1].Reserve[131] := '0';
   Reference[1].Reserve[130] := '0';
   Reference[1].Reserve[129] := '0';
   Reference[1].Reserve[128] := '0';
   Reference[1].Hoist_offset_4[16] := '$00';
   Reference[1].Hoist_offset_4[15] := '$00';
   Reference[1].Hoist_offset_4[14] := '$00';
   Reference[1].Hoist_offset_4[13] := '$00';
   Reference[1].Hoist_offset_4[12] := '$00';
   Reference[1].Hoist_offset_4[11] := '$00';
   Reference[1].Hoist_offset_4[10] := '$00';
   Reference[1].Hoist_offset_4[9] := '$00';
   Reference[1].Hoist_offset_4[8] := '$00';
   Reference[1].Hoist_offset_4[7] := '$00';
   Reference[1].Hoist_offset_4[6] := '$00';
   Reference[1].Hoist_offset_4[5] := '$00';
   Reference[1].Hoist_offset_4[4] := '$00';
   Reference[1].Hoist_offset_4[3] := '$00';
   Reference[1].Hoist_offset_4[2] := '$00';
   Reference[1].Hoist_offset_4[1] := '$00';
   Reference[1].Hoist_offset_3[16] := '$00';
   Reference[1].Hoist_offset_3[15] := '$00';
   Reference[1].Hoist_offset_3[14] := '$00';
   Reference[1].Hoist_offset_3[13] := '$00';
   Reference[1].Hoist_offset_3[12] := '$00';
   Reference[1].Hoist_offset_3[11] := '$00';
   Reference[1].Hoist_offset_3[10] := '$00';
   Reference[1].Hoist_offset_3[9] := '$00';
   Reference[1].Hoist_offset_3[8] := '$00';
   Reference[1].Hoist_offset_3[7] := '$00';
   Reference[1].Hoist_offset_3[6] := '$00';
   Reference[1].Hoist_offset_3[5] := '$00';
   Reference[1].Hoist_offset_3[4] := '$00';
   Reference[1].Hoist_offset_3[3] := '$00';
   Reference[1].Hoist_offset_3[2] := '$00';
   Reference[1].Hoist_offset_3[1] := '$00';
   Reference[1].Hoist_offset_2[16] := '$00';
   Reference[1].Hoist_offset_2[15] := '$00';
   Reference[1].Hoist_offset_2[14] := '$00';
   Reference[1].Hoist_offset_2[13] := '$00';
   Reference[1].Hoist_offset_2[12] := '$00';
   Reference[1].Hoist_offset_2[11] := '$00';
   Reference[1].Hoist_offset_2[10] := '$00';
   Reference[1].Hoist_offset_2[9] := '$00';
   Reference[1].Hoist_offset_2[8] := '$00';
   Reference[1].Hoist_offset_2[7] := '$00';
   Reference[1].Hoist_offset_2[6] := '$00';
   Reference[1].Hoist_offset_2[5] := '$00';
   Reference[1].Hoist_offset_2[4] := '$00';
   Reference[1].Hoist_offset_2[3] := '$00';
   Reference[1].Hoist_offset_2[2] := '$00';
   Reference[1].Hoist_offset_2[1] := '$00';
   Reference[1].Hoist_offset_1[16] := '$00';
   Reference[1].Hoist_offset_1[15] := '$00';
   Reference[1].Hoist_offset_1[14] := '$00';
   Reference[1].Hoist_offset_1[13] := '$00';
   Reference[1].Hoist_offset_1[12] := '$00';
   Reference[1].Hoist_offset_1[11] := '$00';
   Reference[1].Hoist_offset_1[10] := '$00';
   Reference[1].Hoist_offset_1[9] := '$00';
   Reference[1].Hoist_offset_1[8] := '$00';
   Reference[1].Hoist_offset_1[7] := '$00';
   Reference[1].Hoist_offset_1[6] := '$00';
   Reference[1].Hoist_offset_1[5] := '$00';
   Reference[1].Hoist_offset_1[4] := '$00';
   Reference[1].Hoist_offset_1[3] := '$00';
   Reference[1].Hoist_offset_1[2] := '$00';
   Reference[1].Hoist_offset_1[1] := '$00';
   Reference[1].Height[16] := '$00';
   Reference[1].Height[15] := '$00';
   Reference[1].Height[14] := '$00';
   Reference[1].Height[13] := '$00';
   Reference[1].Height[12] := '$00';
   Reference[1].Height[11] := '$00';
   Reference[1].Height[10] := '$00';
   Reference[1].Height[9] := '$00';
   Reference[1].Height[8] := '$00';
   Reference[1].Height[7] := '$00';
   Reference[1].Height[6] := '$00';
   Reference[1].Height[5] := '$00';
   Reference[1].Height[4] := '$00';
   Reference[1].Height[3] := '$00';
   Reference[1].Height[2] := '$00';
   Reference[1].Height[1] := '$00';
   Reference[1].Actionpoint_2[16] := '0';
   Reference[1].Actionpoint_2[15] := '0';
   Reference[1].Actionpoint_2[14] := '0';
   Reference[1].Actionpoint_2[13] := '0';
   Reference[1].Actionpoint_2[12] := '0';
   Reference[1].Actionpoint_2[11] := '0';
   Reference[1].Actionpoint_2[10] := '0';
   Reference[1].Actionpoint_2[9] := '0';
   Reference[1].Actionpoint_2[8] := '0';
   Reference[1].Actionpoint_2[7] := '0';
   Reference[1].Actionpoint_2[6] := '0';
   Reference[1].Actionpoint_2[5] := '0';
   Reference[1].Actionpoint_2[4] := '0';
   Reference[1].Actionpoint_2[3] := '0';
   Reference[1].Actionpoint_2[2] := '0';
   Reference[1].Actionpoint_2[1] := '0';
   Reference[1].Actionpoint_1[16] := '0';
   Reference[1].Actionpoint_1[15] := '0';
   Reference[1].Actionpoint_1[14] := '0';
   Reference[1].Actionpoint_1[13] := '0';
   Reference[1].Actionpoint_1[12] := '0';
   Reference[1].Actionpoint_1[11] := '0';
   Reference[1].Actionpoint_1[10] := '0';
   Reference[1].Actionpoint_1[9] := '0';
   Reference[1].Actionpoint_1[8] := '0';
   Reference[1].Actionpoint_1[7] := '0';
   Reference[1].Actionpoint_1[6] := '0';
   Reference[1].Actionpoint_1[5] := '0';
   Reference[1].Actionpoint_1[4] := '0';
   Reference[1].Actionpoint_1[3] := '0';
   Reference[1].Actionpoint_1[2] := '0';
   Reference[1].Actionpoint_1[1] := '0';
   Reference[1].Sektion[1] := 'b';
   Reference[1].Sektion[2] := 'u';
   Reference[1].Sektion[3] := 'f';
   Reference[1].Sektion[4] := 'f';
   Reference[1].Sektion[5] := 'e';
   Reference[1].Sektion[6] := 'r';
   Reference[1].Sektion[7] := '$00';
   Reference[1].Sektion[8] := '$00';
   Reference[1].Sektion[9] := '$00';
   Reference[1].Sektion[10] := '$00';
   Reference[1].Sektion[11] := '$00';
   Reference[1].Sektion[12] := '$00';
   Reference[1].Sektion[13] := '$00';
   Reference[1].Sektion[14] := '$00';
   Reference[1].Sektion[15] := '$00';
   Reference[1].Sektion[16] := '$00';
   // 19800 more start values not shown
END_DATA_BLOCK

DATA_BLOCK "DB_SDC_TS_REFERENCE_2"   // DB3781
{ S7_Optimized_Access := 'FALSE' }
VERSION : 0.1
   VAR
      HEADER : Struct
         DB_NR : Int := 3781;
         MIN_NR_SEK : Int := 101;
         MAX_NR_SEK : Int := 200;
         START_DAT : Int := 20;
         LAENGE_SEK_DATA : Int := 200;
         Res10 : Int := 0;
         Res12 : Int := 0;
         Res14 : Int := 0;
         Res16 : Int := 0;
         Res18 : Int := 0;
      END_STRUCT;
      Reference : Array[101..200] of Struct
         Sektion : Array[1..16] of Char;
         Actionpoint_1 : Array[1..16] of Char;
         Actionpoint_2 : Array[1..16] of Char;
         Height : Array[1..16] of Char;
         Hoist_offset_1 : Array[1..16] of Char;
         Hoist_offset_2 : Array[1..16] of Char;
         Hoist_offset_3 : Array[1..16] of Char;
         Hoist_offset_4 : Array[1..16] of Char;
         Reserve : Array[128..199] of Char;
      END_STRUCT;
   END_VAR
BEGIN
   Reference[101].Hoist_offset_2[8] := '$00';
   Reference[101].Hoist_offset_2[7] := '$00';
   Reference[101].Hoist_offset_2[6] := '$00';
   Reference[101].Hoist_offset_2[5] := '$00';
   Reference[101].Hoist_offset_2[4] := '$00';
   Reference[101].Hoist_offset_2[3] := '$00';
   Reference[101].Hoist_offset_2[2] := '$00';
   Reference[101].Hoist_offset_2[1] := '$00';
   Reference[101].Hoist_offset_1[16] := '$00';
   Reference[101].Hoist_offset_1[15] := '$00';
   Reference[101].Hoist_offset_1[14] := '$00';
   Reference[101].Hoist_offset_1[13] := '$00';
   Reference[101].Hoist_offset_1[12] := '$00';
   Reference[101].Hoist_offset_1[11] := '$00';
   Reference[101].Hoist_offset_1[10] := '$00';
   Reference[101].Hoist_offset_1[9] := '$00';
   Reference[101].Hoist_offset_1[8] := '$00';
   Reference[101].Hoist_offset_1[7] := '$00';
   Reference[101].Hoist_offset_1[6] := '$00';
   Reference[101].Hoist_offset_1[5] := '$00';
   Reference[101].Hoist_offset_1[4] := '$00';
   Reference[101].Hoist_offset_1[3] := '$00';
   Reference[101].Hoist_offset_1[2] := '$00';
   Reference[101].Hoist_offset_1[1] := '$00';
   Reference[101].Height[16] := '$00';
   Reference[101].Height[15] := '$00';
   Reference[101].Height[14] := '$00';
   Reference[101].Height[13] := '$00';
   Reference[101].Height[12] := '$00';
   Reference[101].Height[11] := '$00';
   Reference[101].Height[10] := '$00';
   Reference[101].Height[9] := '$00';
   Reference[101].Height[8] := '$00';
   Reference[101].Height[7] := '$00';
   Reference[101].Height[6] := '$00';
   Reference[101].Height[5] := '$00';
   Reference[101].Height[4] := '$00';
   Reference[101].Height[3] := '$00';
   Reference[101].Height[2] := '$00';
   Reference[101].Height[1] := '$00';
   Reference[101].Actionpoint_2[16] := '0';
   Reference[101].Actionpoint_2[15] := '0';
   Reference[101].Actionpoint_2[14] := '0';
   Reference[101].Actionpoint_2[13] := '0';
   Reference[101].Actionpoint_2[12] := '0';
   Reference[101].Actionpoint_2[11] := '0';
   Reference[101].Actionpoint_2[10] := '0';
   Reference[101].Actionpoint_2[9] := '0';
   Reference[101].Actionpoint_2[8] := '0';
   Reference[101].Actionpoint_2[7] := '0';
   Reference[101].Actionpoint_2[6] := '0';
   Reference[101].Actionpoint_2[5] := '0';
   Reference[101].Actionpoint_2[4] := '0';
   Reference[101].Actionpoint_2[3] := '0';
   Reference[101].Actionpoint_2[2] := '0';
   Reference[101].Actionpoint_2[1] := '0';
   Reference[101].Actionpoint_1[16] := '0';
   Reference[101].Actionpoint_1[15] := '0';
   Reference[101].Actionpoint_1[14] := '0';
   Reference[101].Actionpoint_1[13] := '0';
   Reference[101].Actionpoint_1[12] := '0';
   Reference[101].Actionpoint_1[11] := '0';
   Reference[101].Actionpoint_1[10] := '0';
   Reference[101].Actionpoint_1[9] := '0';
   Reference[101].Actionpoint_1[8] := '0';
   Reference[101].Actionpoint_1[7] := '0';
   Reference[101].Actionpoint_1[6] := '0';
   Reference[101].Actionpoint_1[5] := '0';
   Reference[101].Actionpoint_1[4] := '0';
   Reference[101].Actionpoint_1[3] := '0';
   Reference[101].Actionpoint_1[2] := '0';
   Reference[101].Actionpoint_1[1] := '0';
   Reference[101].Hoist_offset_3[8] := '$00';
   Reference[101].Hoist_offset_3[7] := '$00';
   Reference[101].Hoist_offset_3[6] := '$00';
   Reference[101].Hoist_offset_3[5] := '$00';
   Reference[101].Hoist_offset_3[4] := '$00';
   Reference[101].Hoist_offset_3[3] := '$00';
   Reference[101].Hoist_offset_3[2] := '$00';
   Reference[101].Hoist_offset_3[1] := '$00';
   Reference[101].Hoist_offset_2[16] := '$00';
   Reference[101].Hoist_offset_2[15] := '$00';
   Reference[101].Hoist_offset_2[14] := '$00';
   Reference[101].Hoist_offset_2[13] := '$00';
   Reference[101].Hoist_offset_2[12] := '$00';
   Reference[101].Hoist_offset_2[11] := '$00';
   Reference[101].Hoist_offset_2[10] := '$00';
   Reference[101].Hoist_offset_2[9] := '$00';
   Reference[101].Hoist_offset_4[8] := '$00';
   Reference[101].Hoist_offset_4[7] := '$00';
   Reference[101].Hoist_offset_4[6] := '$00';
   Reference[101].Hoist_offset_4[5] := '$00';
   Reference[101].Hoist_offset_4[4] := '$00';
   Reference[101].Hoist_offset_4[3] := '$00';
   Reference[101].Hoist_offset_4[2] := '$00';
   Reference[101].Hoist_offset_4[1] := '$00';
   Reference[101].Hoist_offset_3[16] := '$00';
   Reference[101].Hoist_offset_3[15] := '$00';
   Reference[101].Hoist_offset_3[14] := '$00';
   Reference[101].Hoist_offset_3[13] := '$00';
   Reference[101].Hoist_offset_3[12] := '$00';
   Reference[101].Hoist_offset_3[11] := '$00';
   Reference[101].Hoist_offset_3[10] := '$00';
   Reference[101].Hoist_offset_3[9] := '$00';
   Reference[101].Reserve[135] := '0';
   Reference[101].Reserve[134] := '0';
   Reference[101].Reserve[133] := '0';
   Reference[101].Reserve[132] := '0';
   Reference[101].Reserve[131] := '0';
   Reference[101].Reserve[130] := '0';
   Reference[101].Reserve[129] := '0';
   Reference[101].Reserve[128] := '0';
   Reference[101].Hoist_offset_4[16] := '$00';
   Reference[101].Hoist_offset_4[15] := '$00';
   Reference[101].Hoist_offset_4[14] := '$00';
   Reference[101].Hoist_offset_4[13] := '$00';
   Reference[101].Hoist_offset_4[12] := '$00';
   Reference[101].Hoist_offset_4[11] := '$00';
   Reference[101].Hoist_offset_4[10] := '$00';
   Reference[101].Hoist_offset_4[9] := '$00';
   Reference[101].Reserve[151] := ' ';
   Reference[101].Reserve[150] := ' ';
   Reference[101].Reserve[149] := ' ';
   Reference[101].Reserve[148] := ' ';
   Reference[101].Reserve[147] := ' ';
   Reference[101].Reserve[146] := ' ';
   Reference[101].Reserve[145] := ' ';
   Reference[101].Reserve[144] := ' ';
   Reference[101].Reserve[143] := '0';
   Reference[101].Reserve[142] := '0';
   Reference[101].Reserve[141] := '0';
   Reference[101].Reserve[140] := '0';
   Reference[101].Reserve[139] := '0';
   Reference[101].Reserve[138] := '0';
   Reference[101].Reserve[137] := '0';
   Reference[101].Reserve[136] := '0';
   Reference[101].Reserve[167] := ' ';
   Reference[101].Reserve[166] := ' ';
   Reference[101].Reserve[165] := ' ';
   Reference[101].Reserve[164] := ' ';
   Reference[101].Reserve[163] := ' ';
   Reference[101].Reserve[162] := ' ';
   Reference[101].Reserve[161] := ' ';
   Reference[101].Reserve[160] := ' ';
   Reference[101].Reserve[159] := ' ';
   Reference[101].Reserve[158] := ' ';
   Reference[101].Reserve[157] := ' ';
   Reference[101].Reserve[156] := ' ';
   Reference[101].Reserve[155] := ' ';
   Reference[101].Reserve[154] := ' ';
   Reference[101].Reserve[153] := ' ';
   Reference[101].Reserve[152] := ' ';
   Reference[101].Reserve[183] := ' ';
   Reference[101].Reserve[182] := ' ';
   Reference[101].Reserve[181] := ' ';
   Reference[101].Reserve[180] := ' ';
   Reference[101].Reserve[179] := ' ';
   Reference[101].Reserve[178] := ' ';
   Reference[101].Reserve[177] := ' ';
   Reference[101].Reserve[176] := ' ';
   Reference[101].Reserve[175] := ' ';
   Reference[101].Reserve[174] := ' ';
   Reference[101].Reserve[173] := ' ';
   Reference[101].Reserve[172] := ' ';
   Reference[101].Reserve[171] := ' ';
   Reference[101].Reserve[170] := ' ';
   Reference[101].Reserve[169] := ' ';
   Reference[101].Reserve[168] := ' ';
   Reference[101].Reserve[199] := ' ';
   Reference[101].Reserve[198] := ' ';
   Reference[101].Reserve[197] := ' ';
   Reference[101].Reserve[196] := ' ';
   Reference[101].Reserve[195] := ' ';
   Reference[101].Reserve[194] := ' ';
   Reference[101].Reserve[193] := ' ';
   Reference[101].Reserve[192] := ' ';
   Reference[101].Reserve[191] := ' ';
   Reference[101].Reserve[190] := ' ';
   Reference[101].Reserve[189] := ' ';
   Reference[101].Reserve[188] := ' ';
   Reference[101].Reserve[187] := ' ';
   Reference[101].Reserve[186] := ' ';
   Reference[101].Reserve[185] := ' ';
   Reference[101].Reserve[184] := ' ';
   Reference[101].Sektion[1] := ' ';
   Reference[101].Sektion[2] := ' ';
   Reference[101].Sektion[3] := ' ';
   Reference[101].Sektion[4] := ' ';
   Reference[101].Sektion[5] := ' ';
   Reference[101].Sektion[6] := ' ';
   Reference[101].Sektion[7] := ' ';
   Reference[101].Sektion[8] := ' ';
   Reference[101].Sektion[9] := ' ';
   Reference[101].Sektion[10] := ' ';
   Reference[101].Sektion[11] := ' ';
   Reference[101].Sektion[12] := ' ';
   Reference[101].Sektion[13] := ' ';
   Reference[101].Sektion[14] := ' ';
   Reference[101].Sektion[15] := ' ';
   Reference[101].Sektion[16] := ' ';
   // 19800 more start values not shown
END_DATA_BLOCK

